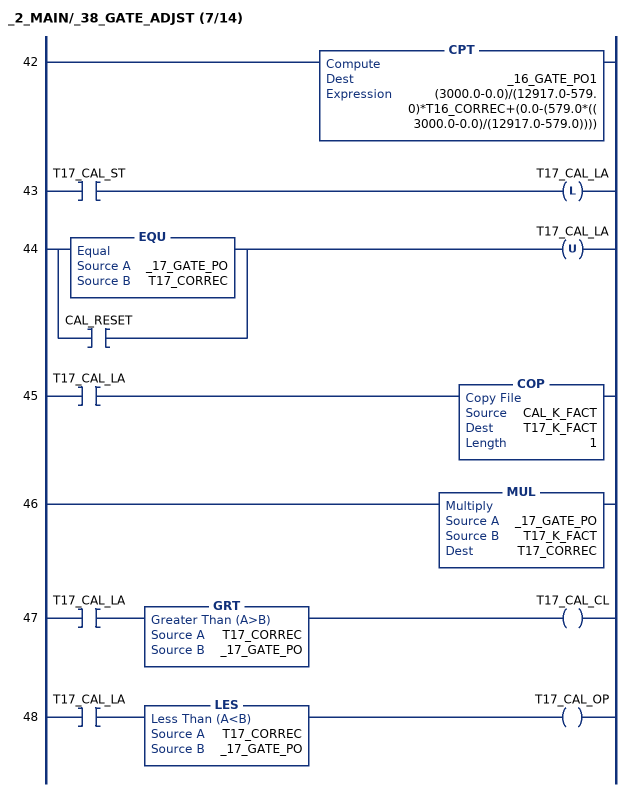
   42: CPT(_16_GATE_PO1,(3000.0-0.0)/(12917.0-579.0)*T16_CORREC+(0.0-(579.0*((3000.0-0.0)/(12917.0-579.0)))));
   43: XIC(T17_CAL_ST)OTL(T17_CAL_LA);
   44: [EQU(_17_GATE_PO,T17_CORREC) ,XIC(CAL_RESET) ]OTU(T17_CAL_LA);
   45: XIC(T17_CAL_LA)COP(CAL_K_FACT,T17_K_FACT,1);
   46: MUL(_17_GATE_PO,T17_K_FACT,T17_CORREC);
   47: XIC(T17_CAL_LA)GRT(T17_CORREC,_17_GATE_PO)OTE(T17_CAL_CL);
   48: XIC(T17_CAL_LA)LES(T17_CORREC,_17_GATE_PO)OTE(T17_CAL_OP);
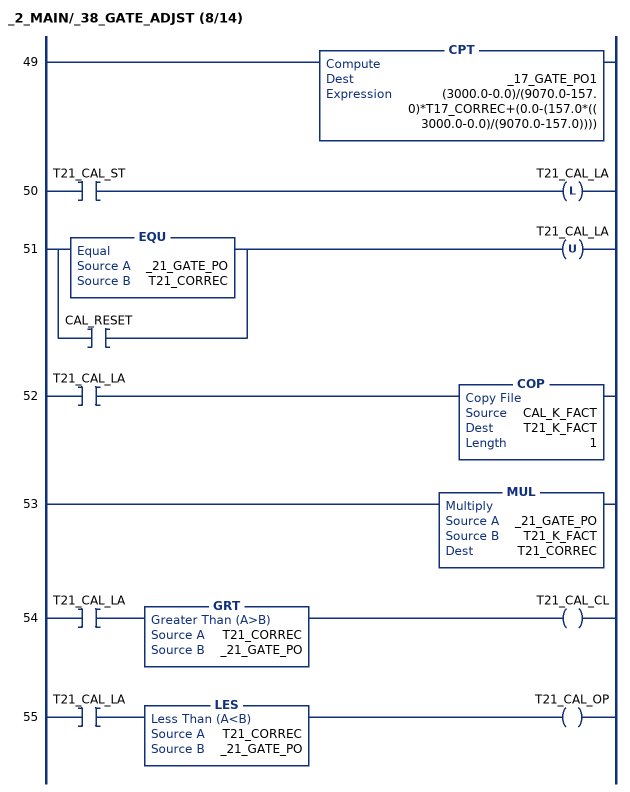
   49: CPT(_17_GATE_PO1,(3000.0-0.0)/(9070.0-157.0)*T17_CORREC+(0.0-(157.0*((3000.0-0.0)/(9070.0-157.0)))));
   50: XIC(T21_CAL_ST)OTL(T21_CAL_LA);
   51: [EQU(_21_GATE_PO,T21_CORREC) ,XIC(CAL_RESET) ]OTU(T21_CAL_LA);
   52: XIC(T21_CAL_LA)COP(CAL_K_FACT,T21_K_FACT,1);
   53: MUL(_21_GATE_PO,T21_K_FACT,T21_CORREC);
   54: XIC(T21_CAL_LA)GRT(T21_CORREC,_21_GATE_PO)OTE(T21_CAL_CL);
   55: XIC(T21_CAL_LA)LES(T21_CORREC,_21_GATE_PO)OTE(T21_CAL_OP);
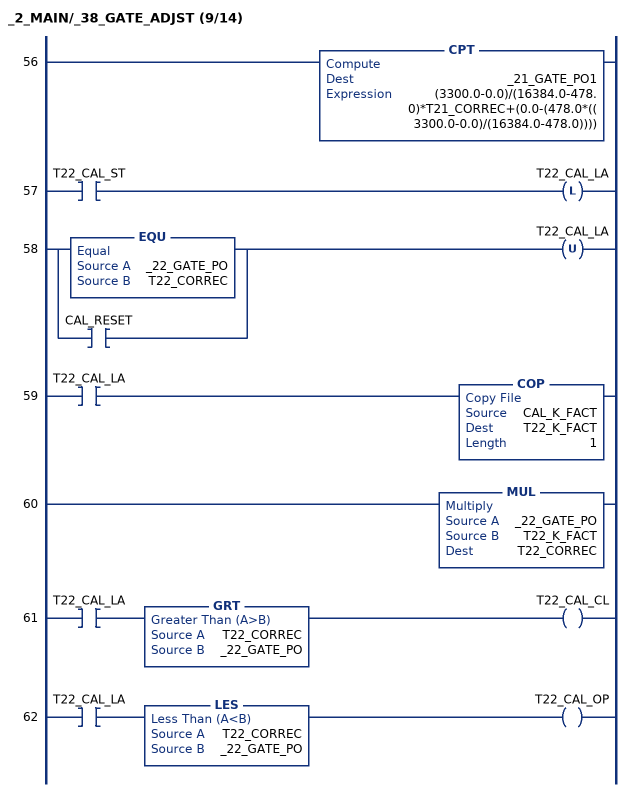
   56: CPT(_21_GATE_PO1,(3300.0-0.0)/(16384.0-478.0)*T21_CORREC+(0.0-(478.0*((3300.0-0.0)/(16384.0-478.0)))));
   57: XIC(T22_CAL_ST)OTL(T22_CAL_LA);
   58: [EQU(_22_GATE_PO,T22_CORREC) ,XIC(CAL_RESET) ]OTU(T22_CAL_LA);
   59: XIC(T22_CAL_LA)COP(CAL_K_FACT,T22_K_FACT,1);
   60: MUL(_22_GATE_PO,T22_K_FACT,T22_CORREC);
   61: XIC(T22_CAL_LA)GRT(T22_CORREC,_22_GATE_PO)OTE(T22_CAL_CL);
   62: XIC(T22_CAL_LA)LES(T22_CORREC,_22_GATE_PO)OTE(T22_CAL_OP);
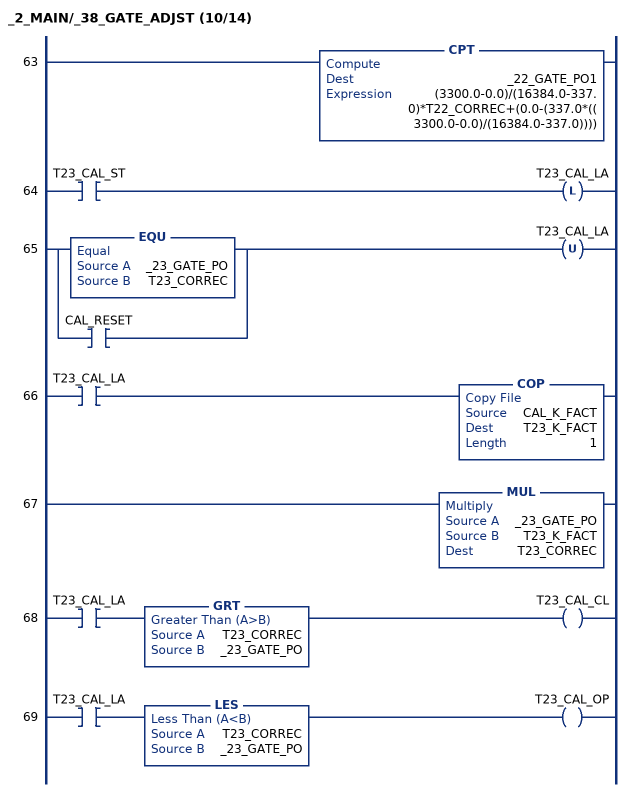
   63: CPT(_22_GATE_PO1,(3300.0-0.0)/(16384.0-337.0)*T22_CORREC+(0.0-(337.0*((3300.0-0.0)/(16384.0-337.0)))));
   64: XIC(T23_CAL_ST)OTL(T23_CAL_LA);
   65: [EQU(_23_GATE_PO,T23_CORREC) ,XIC(CAL_RESET) ]OTU(T23_CAL_LA);
   66: XIC(T23_CAL_LA)COP(CAL_K_FACT,T23_K_FACT,1);
   67: MUL(_23_GATE_PO,T23_K_FACT,T23_CORREC);
   68: XIC(T23_CAL_LA)GRT(T23_CORREC,_23_GATE_PO)OTE(T23_CAL_CL);
   69: XIC(T23_CAL_LA)LES(T23_CORREC,_23_GATE_PO)OTE(T23_CAL_OP);
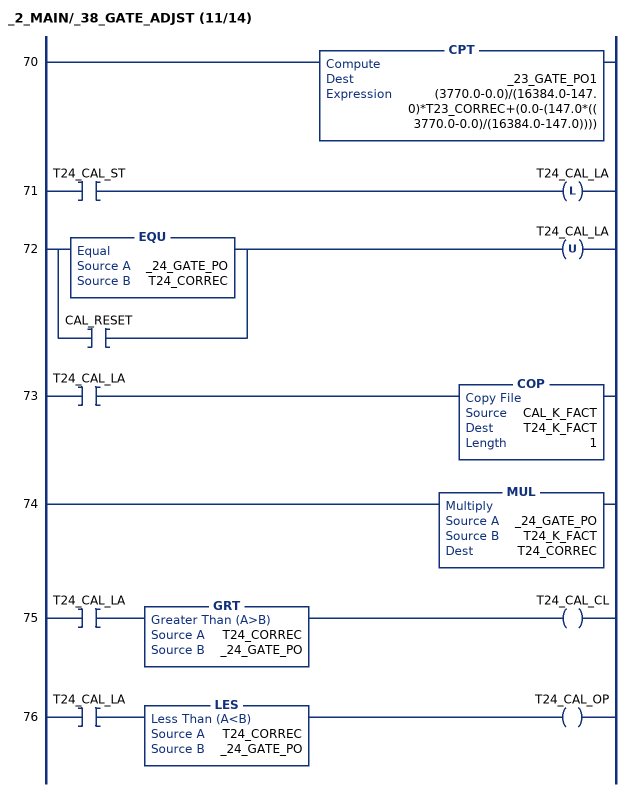
   70: CPT(_23_GATE_PO1,(3770.0-0.0)/(16384.0-147.0)*T23_CORREC+(0.0-(147.0*((3770.0-0.0)/(16384.0-147.0)))));
   71: XIC(T24_CAL_ST)OTL(T24_CAL_LA);
   72: [EQU(_24_GATE_PO,T24_CORREC) ,XIC(CAL_RESET) ]OTU(T24_CAL_LA);
   73: XIC(T24_CAL_LA)COP(CAL_K_FACT,T24_K_FACT,1);
   74: MUL(_24_GATE_PO,T24_K_FACT,T24_CORREC);
   75: XIC(T24_CAL_LA)GRT(T24_CORREC,_24_GATE_PO)OTE(T24_CAL_CL);
   76: XIC(T24_CAL_LA)LES(T24_CORREC,_24_GATE_PO)OTE(T24_CAL_OP);
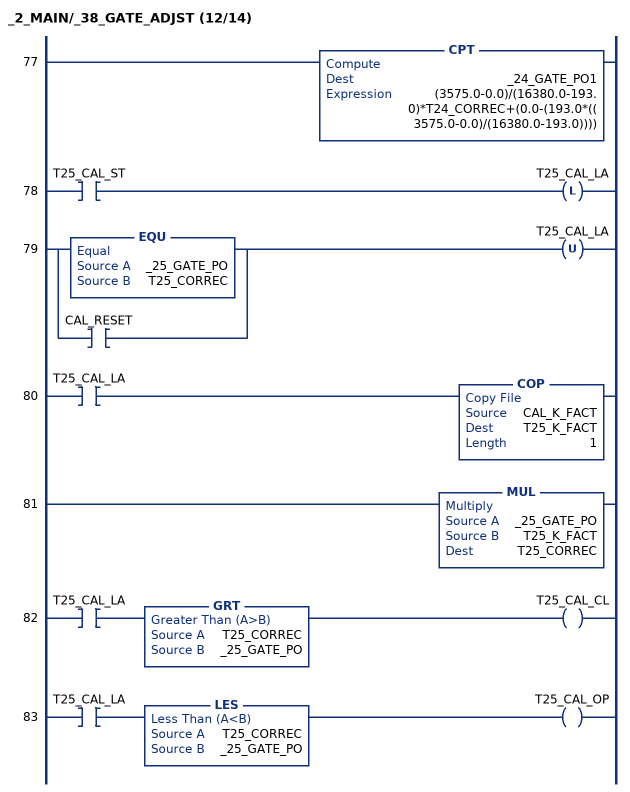
   77: CPT(_24_GATE_PO1,(3575.0-0.0)/(16380.0-193.0)*T24_CORREC+(0.0-(193.0*((3575.0-0.0)/(16380.0-193.0)))));
   78: XIC(T25_CAL_ST)OTL(T25_CAL_LA);
   79: [EQU(_25_GATE_PO,T25_CORREC) ,XIC(CAL_RESET) ]OTU(T25_CAL_LA);
   80: XIC(T25_CAL_LA)COP(CAL_K_FACT,T25_K_FACT,1);
   81: MUL(_25_GATE_PO,T25_K_FACT,T25_CORREC);
   82: XIC(T25_CAL_LA)GRT(T25_CORREC,_25_GATE_PO)OTE(T25_CAL_CL);
   83: XIC(T25_CAL_LA)LES(T25_CORREC,_25_GATE_PO)OTE(T25_CAL_OP);
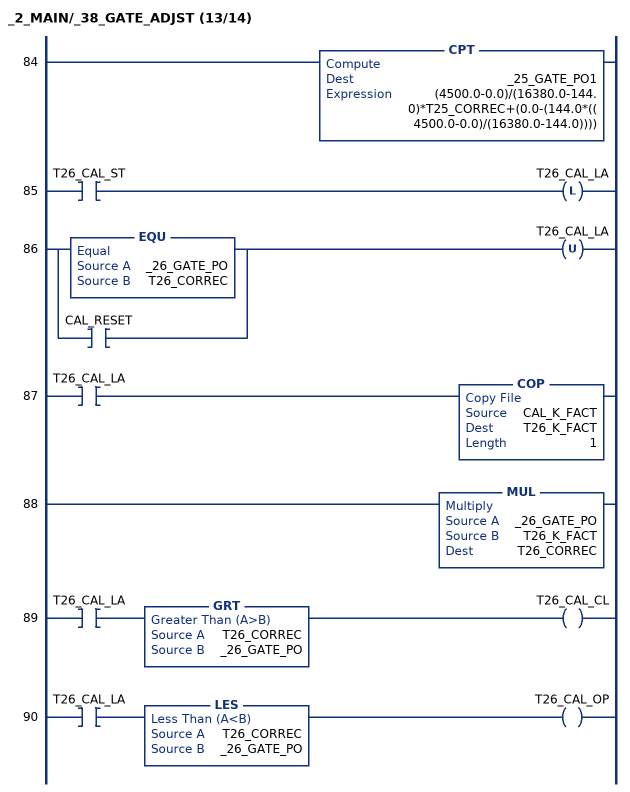
   84: CPT(_25_GATE_PO1,(4500.0-0.0)/(16380.0-144.0)*T25_CORREC+(0.0-(144.0*((4500.0-0.0)/(16380.0-144.0)))));
   85: XIC(T26_CAL_ST)OTL(T26_CAL_LA);
   86: [EQU(_26_GATE_PO,T26_CORREC) ,XIC(CAL_RESET) ]OTU(T26_CAL_LA);
   87: XIC(T26_CAL_LA)COP(CAL_K_FACT,T26_K_FACT,1);
   88: MUL(_26_GATE_PO,T26_K_FACT,T26_CORREC);
   89: XIC(T26_CAL_LA)GRT(T26_CORREC,_26_GATE_PO)OTE(T26_CAL_CL);
   90: XIC(T26_CAL_LA)LES(T26_CORREC,_26_GATE_PO)OTE(T26_CAL_OP);
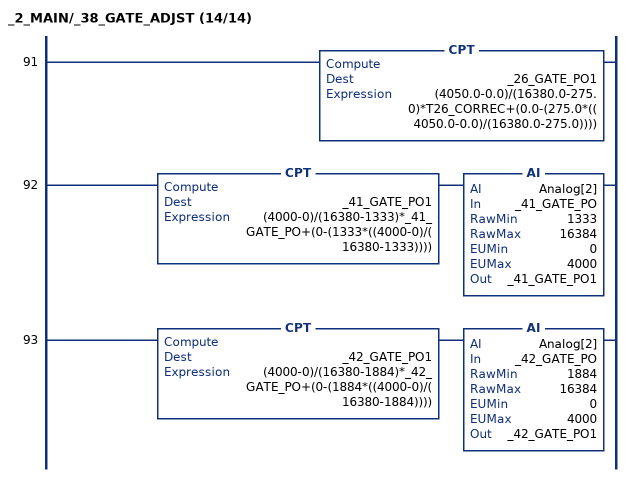
   91: CPT(_26_GATE_PO1,(4050.0-0.0)/(16380.0-275.0)*T26_CORREC+(0.0-(275.0*((4050.0-0.0)/(16380.0-275.0)))));
   92: CPT(_41_GATE_PO1,(4000-0)/(16380-1333)*_41_GATE_PO+(0-(1333*((4000-0)/(16380-1333)))))AI(Analog[2],_41_GATE_PO,1333,16384,0,4000,_41_GATE_PO1);
   93: CPT(_42_GATE_PO1,(4000-0)/(16380-1884)*_42_GATE_PO+(0-(1884*((4000-0)/(16380-1884)))))AI(Analog[2],_42_GATE_PO,1884,16384,0,4000,_42_GATE_PO1);
END_ROUTINE

ROUTINE _39_PUMP_SECUR   (* ladder *)
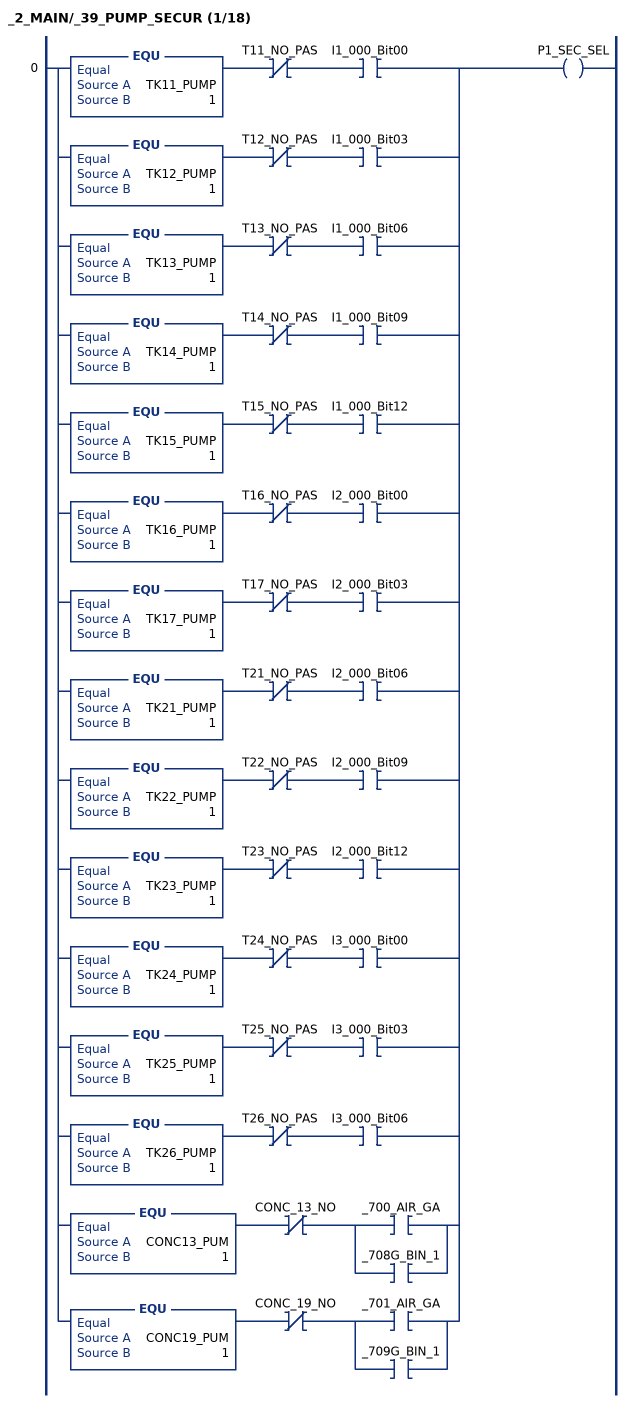
   0: [EQU(TK11_PUMP,1) XIO(T11_NO_PAS) XIC(I1_000_Bit00) ,EQU(TK12_PUMP,1) XIO(T12_NO_PAS) XIC(I1_000_Bit03) ,EQU(TK13_PUMP,1) XIO(T13_NO_PAS) XIC(I1_000_Bit06) ,EQU(TK14_PUMP,1) XIO(T14_NO_PAS) XIC(I1_000_Bit09) ,EQU(TK15_PUMP,1) XIO(T15_NO_PAS) XIC(I1_000_Bit12) ,EQU(TK16_PUMP,1) XIO(T16_NO_PAS) XIC(I2_000_Bit00) ,EQU(TK17_PUMP,1) XIO(T17_NO_PAS) XIC(I2_000_Bit03) ,EQU(TK21_PUMP,1) XIO(T21_NO_PAS) XIC(I2_000_Bit06) ,EQU(TK22_PUMP,1) XIO(T22_NO_PAS) XIC(I2_000_Bit09) ,EQU(TK23_PUMP,1) XIO(T23_NO_PAS) XIC(I2_000_Bit12) ,EQU(TK24_PUMP,1) XIO(T24_NO_PAS) XIC(I3_000_Bit00) ,EQU(TK25_PUMP,1) XIO(T25_NO_PAS) XIC(I3_000_Bit03) ,EQU(TK26_PUMP,1) XIO(T26_NO_PAS) XIC(I3_000_Bit06) ,EQU(CONC13_PUM,1) XIO(CONC_13_NO) [XIC(_700_AIR_GA) ,XIC(_708G_BIN_1) ] ,EQU(CONC19_PUM,1) XIO(CONC_19_NO) [XIC(_701_AIR_GA) ,XIC(_709G_BIN_1) ] ]OTE(P1_SEC_SEL);
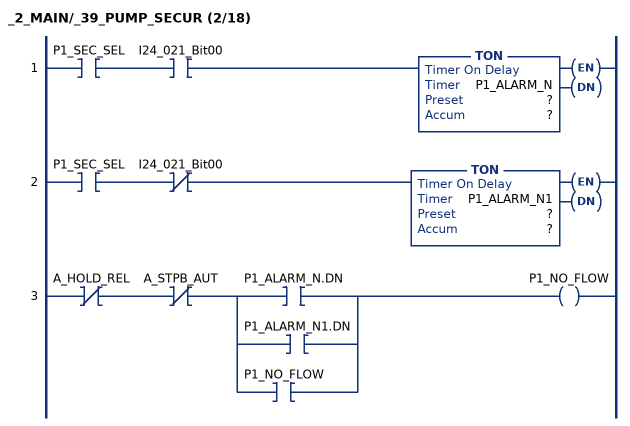
   1: XIC(P1_SEC_SEL)XIC(I24_021_Bit00)TON(P1_ALARM_N,?,?);
   2: XIC(P1_SEC_SEL)XIO(I24_021_Bit00)TON(P1_ALARM_N1,?,?);
   3: XIO(A_HOLD_REL)XIO(A_STPB_AUT)[XIC(P1_ALARM_N.DN) ,XIC(P1_ALARM_N1.DN) ,XIC(P1_NO_FLOW) ]OTE(P1_NO_FLOW);
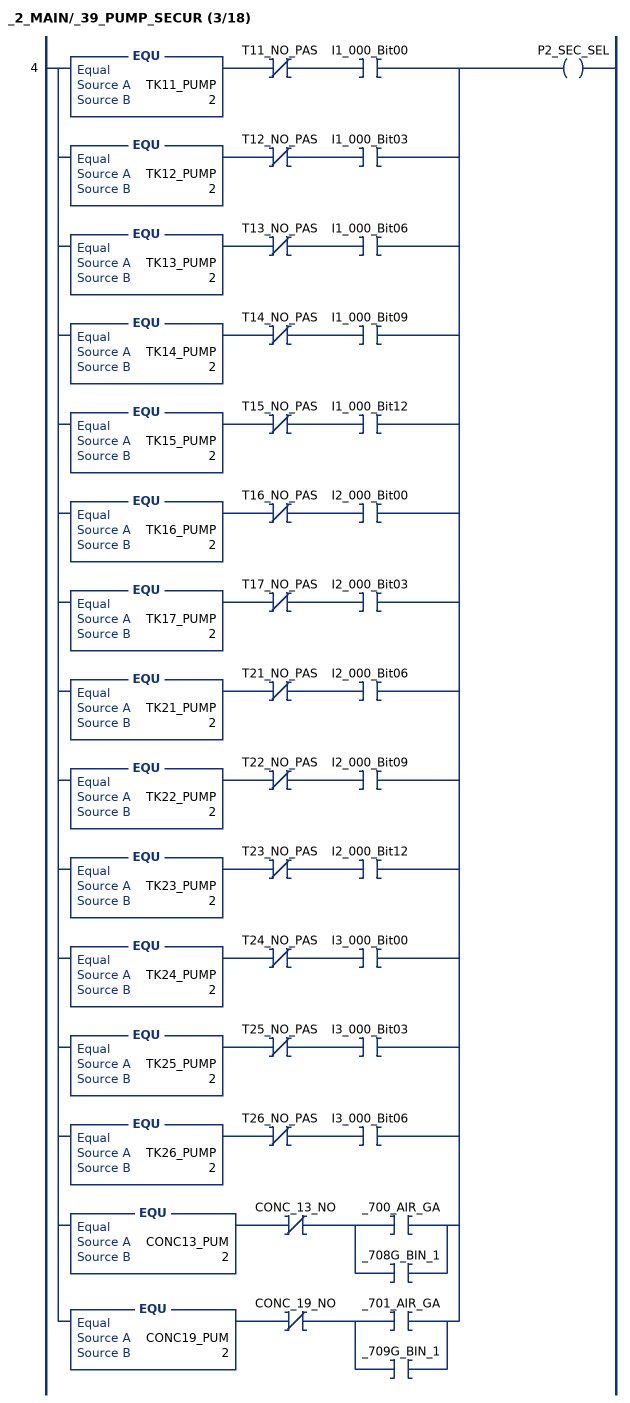
   4: [EQU(TK11_PUMP,2) XIO(T11_NO_PAS) XIC(I1_000_Bit00) ,EQU(TK12_PUMP,2) XIO(T12_NO_PAS) XIC(I1_000_Bit03) ,EQU(TK13_PUMP,2) XIO(T13_NO_PAS) XIC(I1_000_Bit06) ,EQU(TK14_PUMP,2) XIO(T14_NO_PAS) XIC(I1_000_Bit09) ,EQU(TK15_PUMP,2) XIO(T15_NO_PAS) XIC(I1_000_Bit12) ,EQU(TK16_PUMP,2) XIO(T16_NO_PAS) XIC(I2_000_Bit00) ,EQU(TK17_PUMP,2) XIO(T17_NO_PAS) XIC(I2_000_Bit03) ,EQU(TK21_PUMP,2) XIO(T21_NO_PAS) XIC(I2_000_Bit06) ,EQU(TK22_PUMP,2) XIO(T22_NO_PAS) XIC(I2_000_Bit09) ,EQU(TK23_PUMP,2) XIO(T23_NO_PAS) XIC(I2_000_Bit12) ,EQU(TK24_PUMP,2) XIO(T24_NO_PAS) XIC(I3_000_Bit00) ,EQU(TK25_PUMP,2) XIO(T25_NO_PAS) XIC(I3_000_Bit03) ,EQU(TK26_PUMP,2) XIO(T26_NO_PAS) XIC(I3_000_Bit06) ,EQU(CONC13_PUM,2) XIO(CONC_13_NO) [XIC(_700_AIR_GA) ,XIC(_708G_BIN_1) ] ,EQU(CONC19_PUM,2) XIO(CONC_19_NO) [XIC(_701_AIR_GA) ,XIC(_709G_BIN_1) ] ]OTE(P2_SEC_SEL);
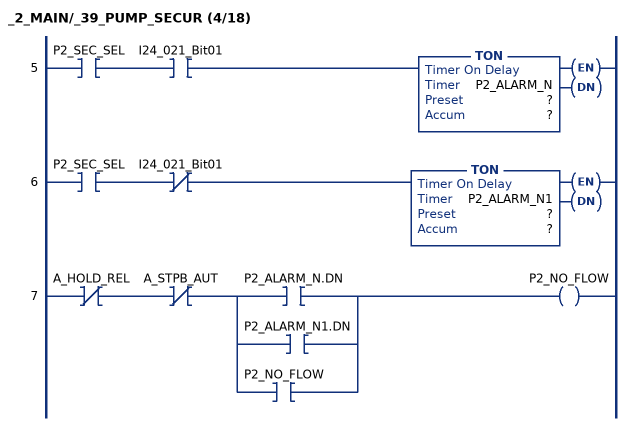
   5: XIC(P2_SEC_SEL)XIC(I24_021_Bit01)TON(P2_ALARM_N,?,?);
   6: XIC(P2_SEC_SEL)XIO(I24_021_Bit01)TON(P2_ALARM_N1,?,?);
   7: XIO(A_HOLD_REL)XIO(A_STPB_AUT)[XIC(P2_ALARM_N.DN) ,XIC(P2_ALARM_N1.DN) ,XIC(P2_NO_FLOW) ]OTE(P2_NO_FLOW);
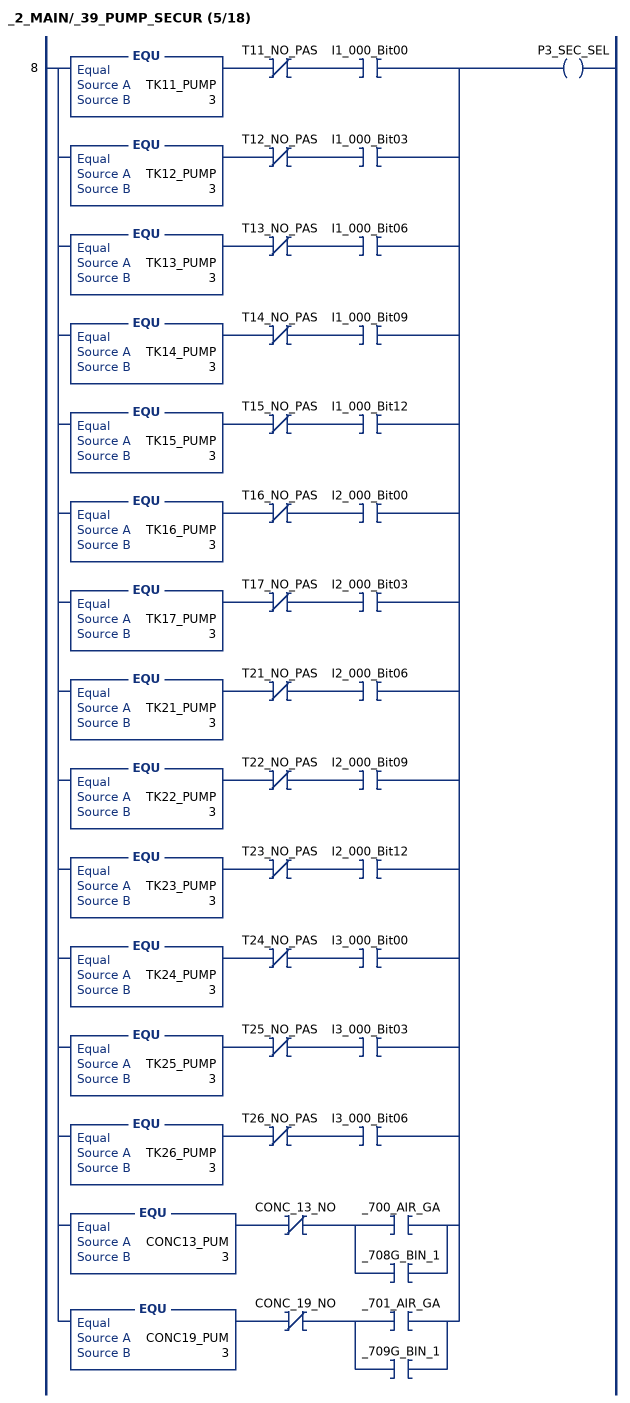
   8: [EQU(TK11_PUMP,3) XIO(T11_NO_PAS) XIC(I1_000_Bit00) ,EQU(TK12_PUMP,3) XIO(T12_NO_PAS) XIC(I1_000_Bit03) ,EQU(TK13_PUMP,3) XIO(T13_NO_PAS) XIC(I1_000_Bit06) ,EQU(TK14_PUMP,3) XIO(T14_NO_PAS) XIC(I1_000_Bit09) ,EQU(TK15_PUMP,3) XIO(T15_NO_PAS) XIC(I1_000_Bit12) ,EQU(TK16_PUMP,3) XIO(T16_NO_PAS) XIC(I2_000_Bit00) ,EQU(TK17_PUMP,3) XIO(T17_NO_PAS) XIC(I2_000_Bit03) ,EQU(TK21_PUMP,3) XIO(T21_NO_PAS) XIC(I2_000_Bit06) ,EQU(TK22_PUMP,3) XIO(T22_NO_PAS) XIC(I2_000_Bit09) ,EQU(TK23_PUMP,3) XIO(T23_NO_PAS) XIC(I2_000_Bit12) ,EQU(TK24_PUMP,3) XIO(T24_NO_PAS) XIC(I3_000_Bit00) ,EQU(TK25_PUMP,3) XIO(T25_NO_PAS) XIC(I3_000_Bit03) ,EQU(TK26_PUMP,3) XIO(T26_NO_PAS) XIC(I3_000_Bit06) ,EQU(CONC13_PUM,3) XIO(CONC_13_NO) [XIC(_700_AIR_GA) ,XIC(_708G_BIN_1) ] ,EQU(CONC19_PUM,3) XIO(CONC_19_NO) [XIC(_701_AIR_GA) ,XIC(_709G_BIN_1) ] ]OTE(P3_SEC_SEL);
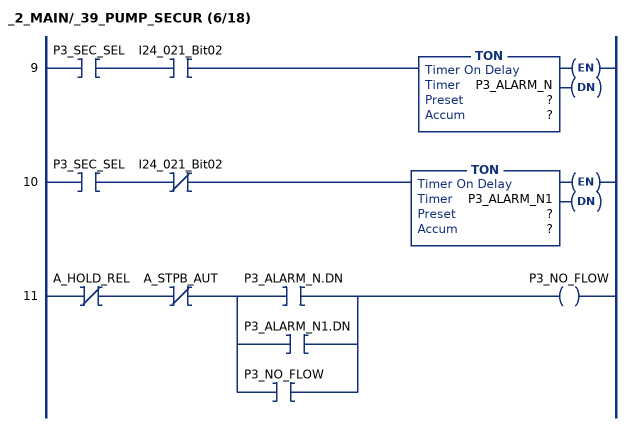
   9: XIC(P3_SEC_SEL)XIC(I24_021_Bit02)TON(P3_ALARM_N,?,?);
   10: XIC(P3_SEC_SEL)XIO(I24_021_Bit02)TON(P3_ALARM_N1,?,?);
   11: XIO(A_HOLD_REL)XIO(A_STPB_AUT)[XIC(P3_ALARM_N.DN) ,XIC(P3_ALARM_N1.DN) ,XIC(P3_NO_FLOW) ]OTE(P3_NO_FLOW);
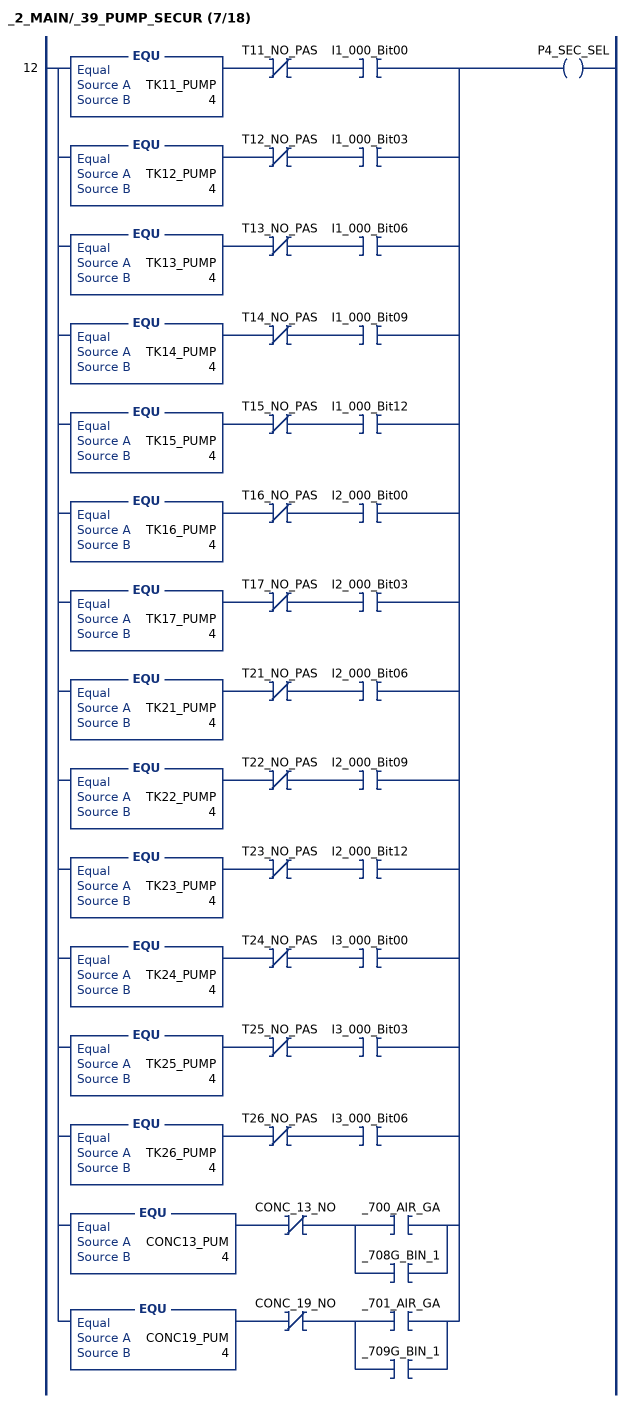
   12: [EQU(TK11_PUMP,4) XIO(T11_NO_PAS) XIC(I1_000_Bit00) ,EQU(TK12_PUMP,4) XIO(T12_NO_PAS) XIC(I1_000_Bit03) ,EQU(TK13_PUMP,4) XIO(T13_NO_PAS) XIC(I1_000_Bit06) ,EQU(TK14_PUMP,4) XIO(T14_NO_PAS) XIC(I1_000_Bit09) ,EQU(TK15_PUMP,4) XIO(T15_NO_PAS) XIC(I1_000_Bit12) ,EQU(TK16_PUMP,4) XIO(T16_NO_PAS) XIC(I2_000_Bit00) ,EQU(TK17_PUMP,4) XIO(T17_NO_PAS) XIC(I2_000_Bit03) ,EQU(TK21_PUMP,4) XIO(T21_NO_PAS) XIC(I2_000_Bit06) ,EQU(TK22_PUMP,4) XIO(T22_NO_PAS) XIC(I2_000_Bit09) ,EQU(TK23_PUMP,4) XIO(T23_NO_PAS) XIC(I2_000_Bit12) ,EQU(TK24_PUMP,4) XIO(T24_NO_PAS) XIC(I3_000_Bit00) ,EQU(TK25_PUMP,4) XIO(T25_NO_PAS) XIC(I3_000_Bit03) ,EQU(TK26_PUMP,4) XIO(T26_NO_PAS) XIC(I3_000_Bit06) ,EQU(CONC13_PUM,4) XIO(CONC_13_NO) [XIC(_700_AIR_GA) ,XIC(_708G_BIN_1) ] ,EQU(CONC19_PUM,4) XIO(CONC_19_NO) [XIC(_701_AIR_GA) ,XIC(_709G_BIN_1) ] ]OTE(P4_SEC_SEL);
